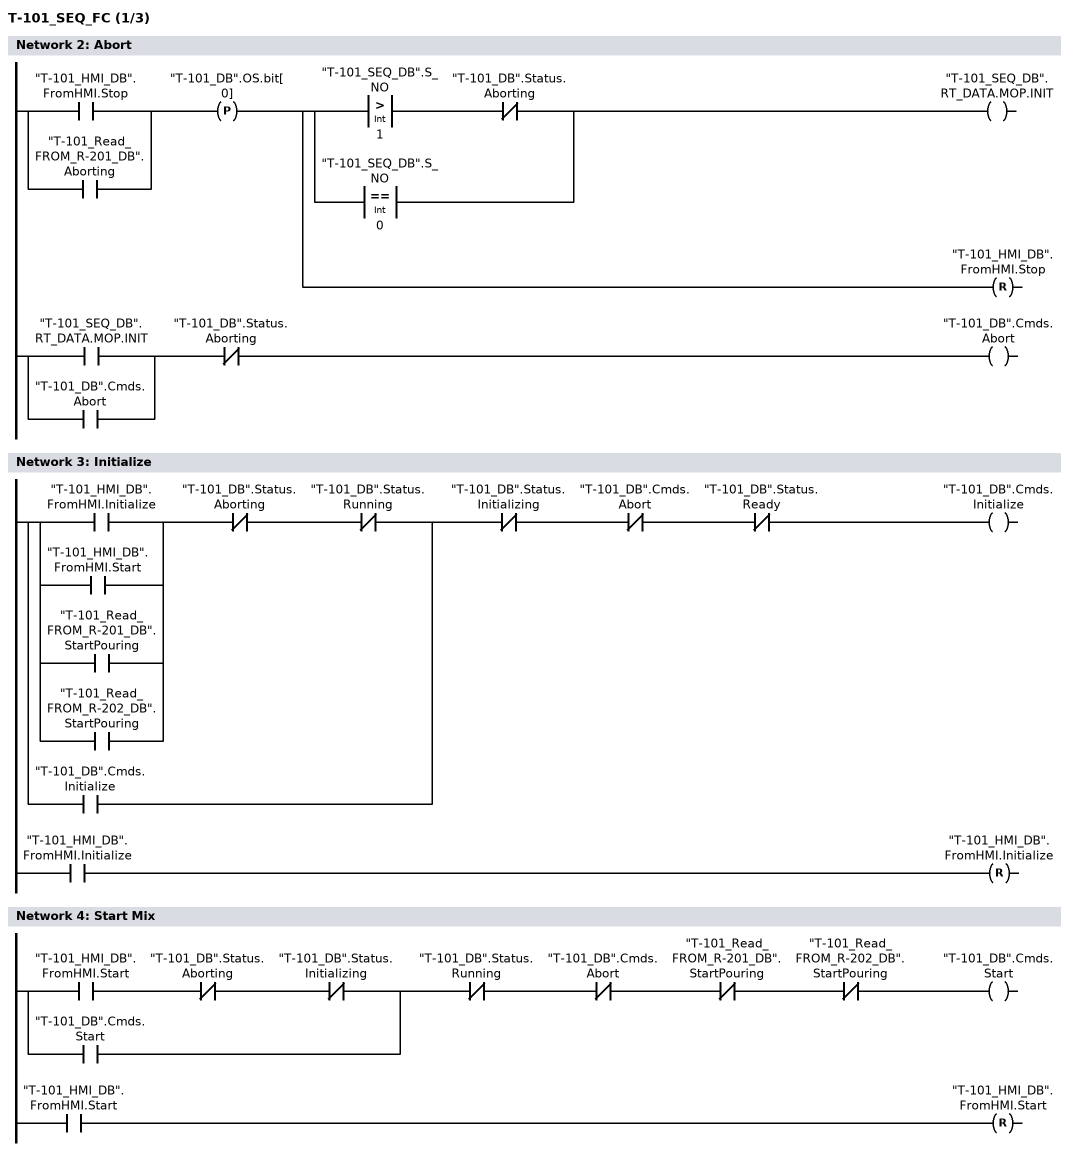
   RUNG wire#powerrail
      Contact( "T-101_HMI_DB".FromHMI.Stop )
      wire#w1
      P_Trig( "T-101_DB".OS.bit[0] )
      wire#w2
      { S7_Templates := "SrcType := Int" } GT_Contact(in1 := "T-101_SEQ_DB".S_NO, in2 := 1)
      I_Contact( "T-101_DB".Status.Aborting )
      wire#w3
      Coil( "T-101_SEQ_DB".RT_DATA.MOP.INIT )
   END_RUNG
   RUNG wire#powerrail
      Contact( "T-101_Read_FROM_R-201_DB".Aborting )
   END_RUNG wire#w1
   RUNG wire#w2
      { S7_Templates := "SrcType := Int" } EQ_Contact(in1 := "T-101_SEQ_DB".S_NO, in2 := 0)
   END_RUNG wire#w3
   RUNG wire#w2
      R_Coil( "T-101_HMI_DB".FromHMI.Stop )
   END_RUNG
   RUNG wire#powerrail
      Contact( "T-101_SEQ_DB".RT_DATA.MOP.INIT )
      wire#w4
      I_Contact( "T-101_DB".Status.Aborting )
      Coil( "T-101_DB".Cmds.Abort )
   END_RUNG
   RUNG wire#powerrail
      Contact( "T-101_DB".Cmds.Abort )
   END_RUNG wire#w4
   // the same network as SCL:
   #_w1 := "T-101_HMI_DB".FromHMI.Stop OR "T-101_Read_FROM_R-201_DB".Aborting;
   #_w2 := #_w1 AND NOT "T-101_DB".OS.bit[0];   // rising edge
   "T-101_DB".OS.bit[0] := #_w1;
   "T-101_SEQ_DB".RT_DATA.MOP.INIT := #_w2 AND ((("T-101_SEQ_DB".S_NO > 1) AND NOT "T-101_DB".Status.Aborting) OR ("T-101_SEQ_DB".S_NO = 0));
   IF #_w2 THEN "T-101_HMI_DB".FromHMI.Stop := FALSE; END_IF;
   "T-101_DB".Cmds.Abort := ("T-101_SEQ_DB".RT_DATA.MOP.INIT OR "T-101_DB".Cmds.Abort) AND NOT "T-101_DB".Status.Aborting;
END_REGION

REGION Network 3: Initialize
   RUNG wire#powerrail
      Contact( "T-101_HMI_DB".FromHMI.Initialize )
      wire#w1
      I_Contact( "T-101_DB".Status.Aborting )
      I_Contact( "T-101_DB".Status.Running )
      wire#w2
      I_Contact( "T-101_DB".Status.Initializing )
      I_Contact( "T-101_DB".Cmds.Abort )
      I_Contact( "T-101_DB".Status.Ready )
      Coil( "T-101_DB".Cmds.Initialize )
   END_RUNG
   RUNG wire#powerrail
      Contact( "T-101_HMI_DB".FromHMI.Start )
   END_RUNG wire#w1
   RUNG wire#powerrail
      Contact( "T-101_Read_FROM_R-201_DB".StartPouring )
   END_RUNG wire#w1
   RUNG wire#powerrail
      Contact( "T-101_Read_FROM_R-202_DB".StartPouring )
   END_RUNG wire#w1
   RUNG wire#powerrail
      Contact( "T-101_DB".Cmds.Initialize )
   END_RUNG wire#w2
   RUNG wire#powerrail
      Contact( "T-101_HMI_DB".FromHMI.Initialize )
      R_Coil( "T-101_HMI_DB".FromHMI.Initialize )
   END_RUNG
   // the same network as SCL:
   "T-101_DB".Cmds.Initialize := ((("T-101_HMI_DB".FromHMI.Initialize OR "T-101_HMI_DB".FromHMI.Start OR "T-101_Read_FROM_R-201_DB".StartPouring OR "T-101_Read_FROM_R-202_DB".StartPouring) AND NOT "T-101_DB".Status.Aborting AND NOT "T-101_DB".Status.Running) OR "T-101_DB".Cmds.Initialize) AND NOT "T-101_DB".Status.Initializing AND NOT "T-101_DB".Cmds.Abort AND NOT "T-101_DB".Status.Ready;
   IF "T-101_HMI_DB".FromHMI.Initialize THEN "T-101_HMI_DB".FromHMI.Initialize := FALSE; END_IF;
END_REGION

REGION Network 4: Start Mix
   RUNG wire#powerrail
      Contact( "T-101_HMI_DB".FromHMI.Start )
      I_Contact( "T-101_DB".Status.Aborting )
      I_Contact( "T-101_DB".Status.Initializing )
      wire#w1
      I_Contact( "T-101_DB".Status.Running )
      I_Contact( "T-101_DB".Cmds.Abort )
      I_Contact( "T-101_Read_FROM_R-201_DB".StartPouring )
      I_Contact( "T-101_Read_FROM_R-202_DB".StartPouring )
      Coil( "T-101_DB".Cmds.Start )
   END_RUNG
   RUNG wire#powerrail
      Contact( "T-101_DB".Cmds.Start )
   END_RUNG wire#w1
   RUNG wire#powerrail
      Contact( "T-101_HMI_DB".FromHMI.Start )
      R_Coil( "T-101_HMI_DB".FromHMI.Start )
   END_RUNG
   // the same network as SCL:
   "T-101_DB".Cmds.Start := (("T-101_HMI_DB".FromHMI.Start AND NOT "T-101_DB".Status.Aborting AND NOT "T-101_DB".Status.Initializing) OR "T-101_DB".Cmds.Start) AND NOT "T-101_DB".Status.Running AND NOT "T-101_DB".Cmds.Abort AND NOT "T-101_Read_FROM_R-201_DB".StartPouring AND NOT "T-101_Read_FROM_R-202_DB".StartPouring;
   IF "T-101_HMI_DB".FromHMI.Start THEN "T-101_HMI_DB".FromHMI.Start := FALSE; END_IF;
END_REGION

REGION Network 5: Procedure Selected
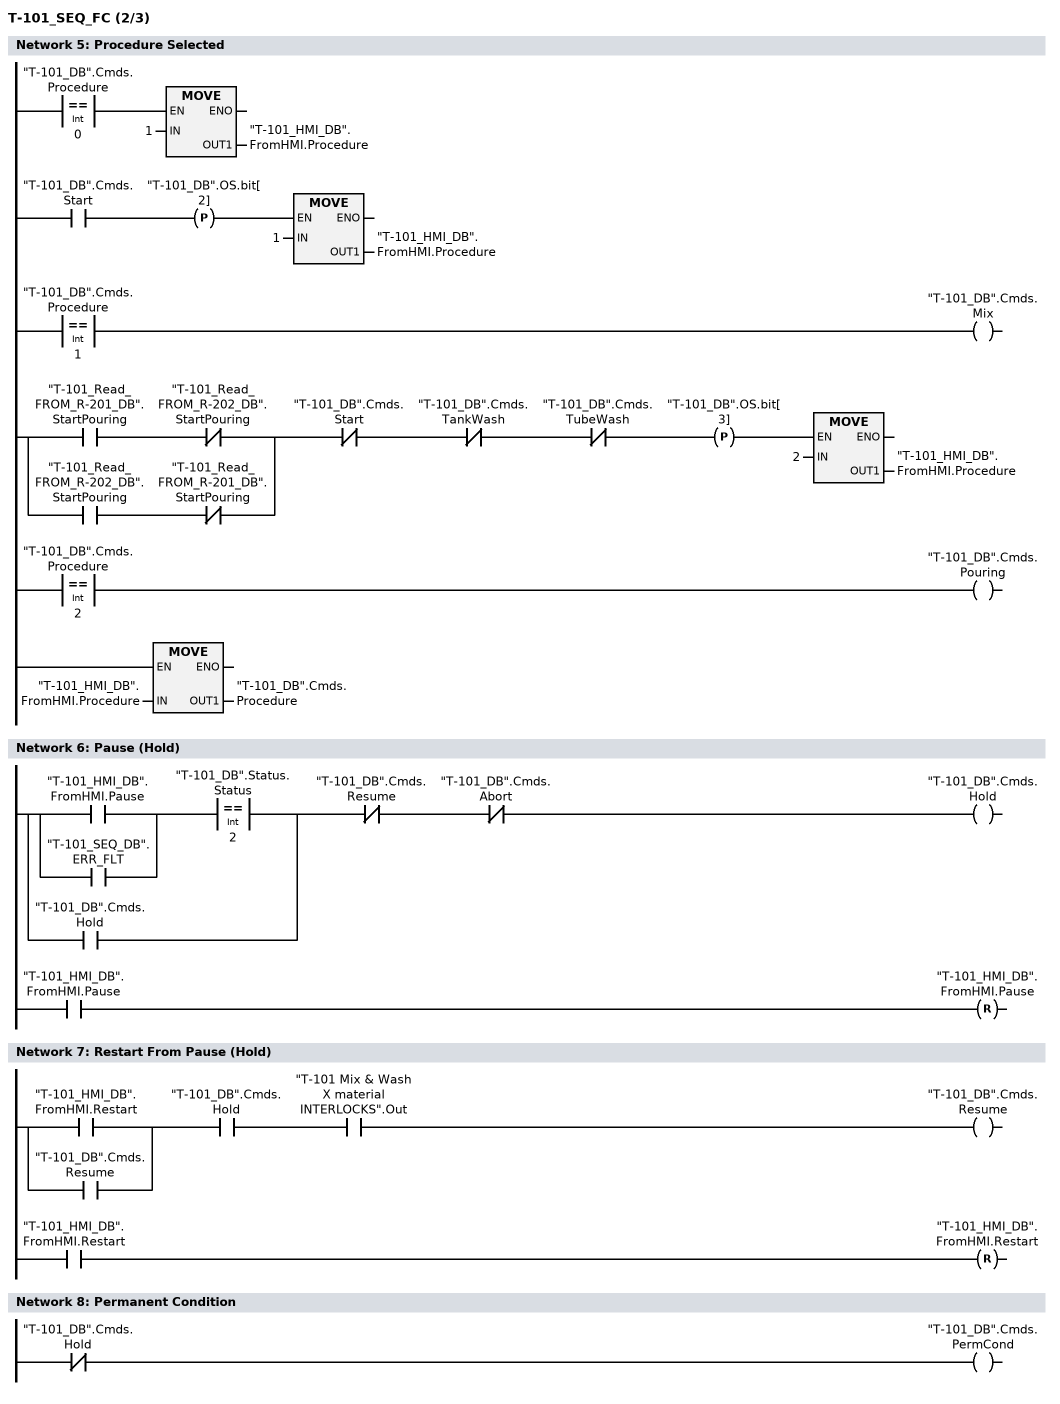
   RUNG wire#powerrail
      { S7_Templates := "SrcType := Int" } EQ_Contact(in1 := "T-101_DB".Cmds.Procedure, in2 := 0)
      Move(in := 1, out1 => "T-101_HMI_DB".FromHMI.Procedure)
   END_RUNG
   RUNG wire#powerrail
      Contact( "T-101_DB".Cmds.Start )
      P_Trig( "T-101_DB".OS.bit[2] )
      Move(in := 1, out1 => "T-101_HMI_DB".FromHMI.Procedure)
   END_RUNG
   RUNG wire#powerrail
      { S7_Templates := "SrcType := Int" } EQ_Contact(in1 := "T-101_DB".Cmds.Procedure, in2 := 1)
      Coil( "T-101_DB".Cmds.Mix )
   END_RUNG
   RUNG wire#powerrail
      Contact( "T-101_Read_FROM_R-201_DB".StartPouring )
      I_Contact( "T-101_Read_FROM_R-202_DB".StartPouring )
      wire#w1
      I_Contact( "T-101_DB".Cmds.Start )
      I_Contact( "T-101_DB".Cmds.TankWash )
      I_Contact( "T-101_DB".Cmds.TubeWash )
      P_Trig( "T-101_DB".OS.bit[3] )
      Move(in := 2, out1 => "T-101_HMI_DB".FromHMI.Procedure)
   END_RUNG
   RUNG wire#powerrail
      Contact( "T-101_Read_FROM_R-202_DB".StartPouring )
      I_Contact( "T-101_Read_FROM_R-201_DB".StartPouring )
   END_RUNG wire#w1
   RUNG wire#powerrail
      { S7_Templates := "SrcType := Int" } EQ_Contact(in1 := "T-101_DB".Cmds.Procedure, in2 := 2)
      Coil( "T-101_DB".Cmds.Pouring )
   END_RUNG
   RUNG wire#powerrail
      Move(in := "T-101_HMI_DB".FromHMI.Procedure, out1 => "T-101_DB".Cmds.Procedure)
   END_RUNG
   // the same network as SCL:
   IF "T-101_DB".Cmds.Procedure = 0 THEN "T-101_HMI_DB".FromHMI.Procedure := 1; END_IF;
   #_w1 := "T-101_DB".Cmds.Start AND NOT "T-101_DB".OS.bit[2];   // rising edge
   "T-101_DB".OS.bit[2] := "T-101_DB".Cmds.Start;
   IF #_w1 THEN "T-101_HMI_DB".FromHMI.Procedure := 1; END_IF;
   "T-101_DB".Cmds.Mix := "T-101_DB".Cmds.Procedure = 1;
   #_w2 := (("T-101_Read_FROM_R-201_DB".StartPouring AND NOT "T-101_Read_FROM_R-202_DB".StartPouring) OR ("T-101_Read_FROM_R-202_DB".StartPouring AND NOT "T-101_Read_FROM_R-201_DB".StartPouring)) AND NOT "T-101_DB".Cmds.Start AND NOT "T-101_DB".Cmds.TankWash AND NOT "T-101_DB".Cmds.TubeWash;
   #_w3 := #_w2 AND NOT "T-101_DB".OS.bit[3];   // rising edge
   "T-101_DB".OS.bit[3] := #_w2;
   IF #_w3 THEN "T-101_HMI_DB".FromHMI.Procedure := 2; END_IF;
   "T-101_DB".Cmds.Pouring := "T-101_DB".Cmds.Procedure = 2;
   "T-101_DB".Cmds.Procedure := "T-101_HMI_DB".FromHMI.Procedure;
END_REGION

REGION Network 6: Pause (Hold)
   RUNG wire#powerrail
      Contact( "T-101_HMI_DB".FromHMI.Pause )
      wire#w1
      { S7_Templates := "SrcType := Int" } EQ_Contact(in1 := "T-101_DB".Status.Status, in2 := 2)
      wire#w2
      I_Contact( "T-101_DB".Cmds.Resume )
      I_Contact( "T-101_DB".Cmds.Abort )
      Coil( "T-101_DB".Cmds.Hold )
   END_RUNG
   RUNG wire#powerrail
      Contact( "T-101_SEQ_DB".ERR_FLT )
   END_RUNG wire#w1
   RUNG wire#powerrail
      Contact( "T-101_DB".Cmds.Hold )
   END_RUNG wire#w2
   RUNG wire#powerrail
      Contact( "T-101_HMI_DB".FromHMI.Pause )
      R_Coil( "T-101_HMI_DB".FromHMI.Pause )
   END_RUNG
   // the same network as SCL:
   "T-101_DB".Cmds.Hold := ((("T-101_HMI_DB".FromHMI.Pause OR "T-101_SEQ_DB".ERR_FLT) AND ("T-101_DB".Status.Status = 2)) OR "T-101_DB".Cmds.Hold) AND NOT "T-101_DB".Cmds.Resume AND NOT "T-101_DB".Cmds.Abort;
   IF "T-101_HMI_DB".FromHMI.Pause THEN "T-101_HMI_DB".FromHMI.Pause := FALSE; END_IF;
END_REGION

REGION Network 7: Restart From Pause (Hold)
   RUNG wire#powerrail
      Contact( "T-101_HMI_DB".FromHMI.Restart )
      wire#w1
      Contact( "T-101_DB".Cmds.Hold )
      Contact( "T-101 Mix & Wash X material INTERLOCKS".Out )
      Coil( "T-101_DB".Cmds.Resume )
   END_RUNG
   RUNG wire#powerrail
      Contact( "T-101_DB".Cmds.Resume )
   END_RUNG wire#w1
   RUNG wire#powerrail
      Contact( "T-101_HMI_DB".FromHMI.Restart )
      R_Coil( "T-101_HMI_DB".FromHMI.Restart )
   END_RUNG
   // the same network as SCL:
   "T-101_DB".Cmds.Resume := ("T-101_HMI_DB".FromHMI.Restart OR "T-101_DB".Cmds.Resume) AND "T-101_DB".Cmds.Hold AND "T-101 Mix & Wash X material INTERLOCKS".Out;
   IF "T-101_HMI_DB".FromHMI.Restart THEN "T-101_HMI_DB".FromHMI.Restart := FALSE; END_IF;
END_REGION

REGION Network 8: Permanent Condition
   RUNG wire#powerrail
      I_Contact( "T-101_DB".Cmds.Hold )
      Coil( "T-101_DB".Cmds.PermCond )
   END_RUNG
   // the same network as SCL:
   "T-101_DB".Cmds.PermCond := NOT "T-101_DB".Cmds.Hold;
END_REGION

REGION Network 9: Tank Wash
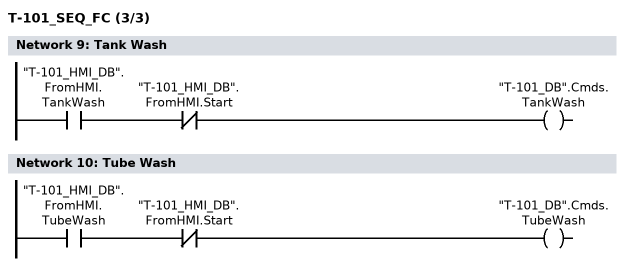
   RUNG wire#powerrail
      Contact( "T-101_HMI_DB".FromHMI.TankWash )
      I_Contact( "T-101_HMI_DB".FromHMI.Start )
      Coil( "T-101_DB".Cmds.TankWash )
   END_RUNG
   // the same network as SCL:
   "T-101_DB".Cmds.TankWash := "T-101_HMI_DB".FromHMI.TankWash AND NOT "T-101_HMI_DB".FromHMI.Start;
END_REGION

REGION Network 10: Tube Wash
   RUNG wire#powerrail
      Contact( "T-101_HMI_DB".FromHMI.TubeWash )
      I_Contact( "T-101_HMI_DB".FromHMI.Start )
      Coil( "T-101_DB".Cmds.TubeWash )
   END_RUNG
   // the same network as SCL:
   "T-101_DB".Cmds.TubeWash := "T-101_HMI_DB".FromHMI.TubeWash AND NOT "T-101_HMI_DB".FromHMI.Start;
END_REGION

REGION Network 11 (SCL): Sequence Status
   IF "T-101_SEQ_DB".S_NO = 1 THEN
       "T-101_DB".Status.Status := 1; //Idle
   ELSIF ("T-101_SEQ_DB".S_NO > 1 AND "T-101_SEQ_DB".S_NO < 150) AND NOT "T-101_SEQ_DB".ERR_FLT AND NOT "T-101_DB".Cmds.Hold THEN
       "T-101_DB".Status.Status := 2; //Running
   ELSIF "T-101_SEQ_DB".S_NO >= 151 AND "T-101_SEQ_DB".S_NO <= 160 AND NOT "T-101_SEQ_DB".ERR_FLT THEN
       "T-101_DB".Status.Status := 3; // Stopping
   ELSIF "T-101_SEQ_DB".ERR_FLT AND ("T-101_SEQ_DB".S_NO > 1 AND "T-101_SEQ_DB".S_NO < 150) THEN
       "T-101_DB".Status.Status := 4; // Held
   ELSIF "T-101_SEQ_DB".ERR_FLT AND ("T-101_SEQ_DB".S_NO > 1 AND "T-101_SEQ_DB".S_NO < 150) AND "T-101_Aux_DB"."Bool".TOff THEN
       "T-101_DB".Status.Status := 5; // Holding
   ELSE
       "T-101_DB".Status.Status := 6; // Unknown
   END_IF;

   "T-101_DB".Status.Running := ("T-101_SEQ_DB".S_NO > 3 AND "T-101_SEQ_DB".S_NO <= 150);
   "T-101_DB".Status.Initializing := ("T-101_SEQ_DB".S_NO >= 141 AND "T-101_SEQ_DB".S_NO <= 150);
   //"T-101_DB".Status.Aborting := ("T-101_SEQ_DB".S_NO >= 151 AND "T-101_SEQ_DB".S_NO <= 160);

   //Enable/Disable HMI Start/Stop Button
   "T-101_HMI_DB".ToHMI.EnStopButton := ("T-101_DB".Status.Status > 1) OR "T-101_DB".Status.Step = 0; //Enable HMI Stop Button
   "T-101_HMI_DB".ToHMI.EnStartButton := "T-101_DB".Status.Status = 1; //Idle
   "T-101_HMI_DB".ToHMI.EnPauseButton := "T-101_DB".Status.Status = 2; //Enable Pause Button
   "T-101_HMI_DB".ToHMI.EnRestartButton :=  "T-101_DB".Status.Status = 4 ; //Enable Restart Button

   //****Interlock Activated
   "T-101_HMI_DB".ToHMI.InterlockActivated := "T-101 Mix & Wash X material INTERLOCKS".Out;
END_REGION

REGION Network 12 (SCL): Sequence Step
   "T-101_DB".Status.Step := "T-101_SEQ_DB".S_NO;
END_REGION

REGION Network 13 (SCL): Sequence state (Procedure running)
   IF "T-101_SEQ_DB".S_NO = 3 OR "T-101_SEQ_DB".S_NO = 4 THEN
       "T-101_DB".Status.State := 1; //Ready
   ELSIF "T-101_SEQ_DB".S_NO >= 21 AND "T-101_SEQ_DB".S_NO <= 60 THEN
       "T-101_DB".Status.State := 2; //Mixing 
   ELSIF "T-101_SEQ_DB".S_NO >= 61 AND "T-101_SEQ_DB".S_NO <= 80 THEN
       "T-101_DB".Status.State := 3; //Pouring
   ELSIF "T-101_SEQ_DB".S_NO >= 141 AND "T-101_SEQ_DB".S_NO <= 150 THEN
       "T-101_DB".Status.State := 4; //Initializing
   ELSIF "T-101_SEQ_DB".S_NO >= 151 AND "T-101_SEQ_DB".S_NO <= 160 THEN
       "T-101_DB".Status.State := 5; //Aborting
   ELSE
       "T-101_DB".Status.State := 0;
   END_IF;
END_REGION

REGION Network 14: Sequence State
END_REGION
END_FUNCTION

FUNCTION "T-101_FC_Outputs" : Void   // FC81, SCL
{ S7_Optimized_Access := 'TRUE' }
VERSION : 0.1
   VAR_TEMP
      Pump_A : Struct
         Cond_01 : Bool;   // Condition 01
         Cond_02 : Bool;
         Cond_03 : Bool;   // Condition 03
      END_STRUCT;
      Pump_B : Struct
         Cond_01 : Bool;   // Condition 01
         Cond_02 : Bool;   // Condition 02
         Cond_03 : Bool;   // Condition 03
      END_STRUCT;
      XV : Struct
         "1011" : Bool;
         "1041" : Bool;
         "1013" : Bool;
      END_STRUCT;
      RouteOpened : Bool;
      PumpsOff : Bool;
      Recirculating : Bool;
   END_VAR
BEGIN
   //****** Equipmens Activation*******
   //
   //**************************************************************
   //

   //
   //IF "AlwaysFALSE" THEN
       //***********************************************Tank Outlet Valve**********************************************************************
       IF  "XV-1011_DB".Mode=0 THEN
           "T-101_DB".Equipments.Valves."XV-1011".CmdOn := "T-101_DB".Equipments.Valves."XV-1011".Enable AND NOT "T-101_DB".Cmds.Hold;
           //Delay Off To avoid Overpressure the Lines
           #XV."1011" := "T-101_DB".Equipments.Valves."XV-1011".CmdOn;
           "T-101_Aux_DB".Timer."XV-1011".TOF(IN := #XV."1011",
                                              PT := "T-101_Aux_DB".Constants.CmdDelay);
           //Command to the Valve
           IF "T-101_Aux_DB".Timer."XV-1011".Q THEN
               "XV-1011_DB".CMD := 2;
           ELSE
               "XV-1011_DB".CMD := 1;
           END_IF;
           "T-101_DB".Equipments.Valves."XV-1011".TurningOff := NOT "T-101_DB".Equipments.Valves."XV-1011".CmdOn AND "T-101_Aux_DB".Timer."XV-1011".Q;
       END_IF;
       //***********************************************Tank Inlet Valve**********************************************************************
       IF  "XV-1041_DB".Mode = 0 THEN
           "T-101_DB".Equipments.Valves."XV-1041".CmdOn := "T-101_DB".Equipments.Valves."XV-1041".Enable AND NOT "T-101_DB".Cmds.Hold;
           //Delay Off To avoid Overpressure the Lines
           #XV."1041" := "T-101_DB".Equipments.Valves."XV-1041".CmdOn;
           "T-101_Aux_DB".Timer."XV-1041".TOF(IN := #XV."1041",
                                              PT := "T-101_Aux_DB".Constants.CmdDelay);
           //Command to the Valve
           IF "T-101_Aux_DB".Timer."XV-1041".Q THEN
               "XV-1041_DB".CMD := 2;
           ELSE
               "XV-1041_DB".CMD := 1;
           END_IF;
           "T-101_DB".Equipments.Valves."XV-1041".TurningOff := NOT "T-101_DB".Equipments.Valves."XV-1041".CmdOn AND "T-101_Aux_DB".Timer."XV-1041".Q;
       END_IF;
       //***********************************************Tank Transfer Valve**********************************************************************
       IF  "XV-1013_DB".Mode = 0 THEN
           "T-101_DB".Equipments.Valves."XV-1013".CmdOn := "T-101_DB".Equipments.Valves."XV-1013".Enable AND NOT "T-101_DB".Cmds.Hold;
           //Delay Off To avoid Overpressure the Lines
           #XV."1013" := "T-101_DB".Equipments.Valves."XV-1013".CmdOn;
           "T-101_Aux_DB".Timer."XV-1013".TOF(IN := #XV."1013",
                                              PT := "T-101_Aux_DB".Constants.CmdDelay);
           //Command to the Valve
           IF "T-101_Aux_DB".Timer."XV-1013".Q THEN
               "XV-1013_DB".CMD := 2;
           ELSE
               "XV-1013_DB".CMD := 1;
           END_IF;
           "T-101_DB".Equipments.Valves."XV-1013".TurningOff := NOT "T-101_DB".Equipments.Valves."XV-1013".CmdOn AND "T-101_Aux_DB".Timer."XV-1013".Q;
       END_IF;
      // IF NOT "TestDB".DesablePmps_T101 THEN
           //***********************************************Feed Water Pump A**********************************************************************
           // Condition to CmdOn "On Command" 
           IF  "P-101A_DB".Config.HMI.Enable_HMI_Controls=1 THEN
               #Pump_A.Cond_01 := "T-101_DB".Equipments.Pumps."P-101A".Enable AND ("T-101_DB".PmpSel."P-101AB" = 1 OR "T-101_DB".PmpSel."P-101AB" = 3);
               #Pump_A.Cond_02 := "T-101_Write_TO_R-201_DB".RouteOpened AND "T-101_Read_FROM_R-201_DB".RouteOpened OR ("T-101_Write_TO_R-202_DB".RouteOpened AND "T-101_Read_FROM_R-202_DB".RouteOpened); //Route Open to sent to the Reactor
               #Pump_A.Cond_03 := "XV-1011_DB".OS AND "XV-1013_DB".CS; //Route open to Recirculate
               "T-101_DB".Equipments.Pumps."P-101A".CmdOn := #Pump_A.Cond_01 AND (#Pump_A.Cond_02 OR #Pump_A.Cond_03) AND NOT "T-101_DB".Cmds.Hold;
               IF "T-101_DB".Equipments.Pumps."P-101A".CmdOn THEN
                   "P-101A_DB".Stop_CMD := False;
                   "P-101A_DB".Start_CMD := true;
                   "P-101A_DB".ON := TRUE;
                   "P-101A_DB".OFF := FALSE;
               ELSE
                   "P-101A_DB".Stop_CMD := true;
                   "P-101A_DB".Start_CMD :=false;
                   "P-101A_DB".ON := FALSE;
                   "P-101A_DB".OFF := TRUE;
               END_IF;
           END_IF;
           //***********************************************Feed Water Pump B**********************************************************************
           // Condition to CmdOn "On Command" 
           IF  "P-101B_DB".Config.HMI.Enable_HMI_Controls = 1 THEN
               #Pump_B.Cond_01 := "T-101_DB".Equipments.Pumps."P-101B".Enable AND ("T-101_DB".PmpSel."P-101AB" = 2 OR "T-101_DB".PmpSel."P-101AB" = 3);
               #Pump_B.Cond_02 := "T-101_Write_TO_R-201_DB".RouteOpened AND "T-101_Read_FROM_R-201_DB".RouteOpened  OR ("T-101_Write_TO_R-202_DB".RouteOpened AND "T-101_Read_FROM_R-202_DB".RouteOpened); //Route Open to sent to the Reactor
               #Pump_B.Cond_03 := "XV-1011_DB".OS AND "XV-1013_DB".CS; //Route open to Recirculate
               "T-101_DB".Equipments.Pumps."P-101B".CmdOn := #Pump_B.Cond_01 AND (#Pump_B.Cond_02 OR #Pump_B.Cond_03) AND NOT "T-101_DB".Cmds.Hold;
               IF "T-101_DB".Equipments.Pumps."P-101B".CmdOn THEN
                   "P-101B_DB".Stop_CMD := False;
                   "P-101B_DB".Start_CMD := true;
                   "P-101B_DB".ON := TRUE;
                   "P-101B_DB".OFF := FALSE;
               ELSE
                   "P-101B_DB".Stop_CMD := True;
                   "P-101B_DB".Start_CMD := False;
                   "P-101B_DB".ON := FALSE;
                   "P-101B_DB".OFF := TRUE;
               END_IF;
           END_IF;
       //END_IF;
           //***********************************************Mixer***********************************************************************
           IF "VFD-T101A_DB".HMI.Controls.Mode = 2 THEN
               "T-101_DB".Equipments.VFD."VFD-1011".CmdOn := "T-101_DB".Equipments.VFD."VFD-1011".Enable AND NOT "T-101_DB".Cmds.Hold;
               IF "T-101_DB".Equipments.VFD."VFD-1011".CmdOn THEN
                   "VFD-T101A_DB".PLCCommand := TRUE;
               ELSE
                   "VFD-T101A_DB".PLCCommand := FALSE;
               END_IF;
           END_IF;
       //END_IF;


   //END_IF;

   //***************Interlocks to R-201***************//
   //*****Recirculating*****//
   #Recirculating := ("P-101A_DB".CF OR "P-101B_DB".CF) AND ("XV-1011_DB".OS AND "XV-1013_DB".CS) AND ("FT-1011_DB".SAI > 0.2);

   "T-101_Write_TO_R-201_DB".Recirculating :=    #Recirculating;
   "T-101_Write_TO_R-202_DB".Recirculating :=    #Recirculating;
   //****Route open to R-201*****//
           #RouteOpened := "XV-1011_DB".OS AND "XV-1013_DB".OS;

   "T-101_Write_TO_R-201_DB".RouteOpened :=   #RouteOpened ;
   "T-101_Write_TO_R-202_DB".RouteOpened := #RouteOpened;
   //*****Pumps OFF*****//
   #PumpsOff := NOT "P-101A_DB".CF AND NOT "P-101B_DB".CF AND ("PT-101A_DB".SAI < 0.8 AND "PT-101B_DB".SAI < 0.8);

   "T-101_Write_TO_R-201_DB".PupmsOFF :=  #PumpsOff ;
   "T-101_Write_TO_R-202_DB".PupmsOFF :=  #PumpsOff ;

           //********************Tank Internal Status*********************************
   "T-101_DB".Status.PouringRunning := ("T-101_DB".Status.Step = 61 OR "T-101_DB".Status.Step = 62 OR "T-101_DB".Status.Step = 63) AND (#RouteOpened AND NOT #PumpsOff);

   //***************Interlocks to T-104***************//
   "T-101_Write_TO_T-104_DB".ReqWaterToMix := "XV-1041_DB".OS AND "T-101_DB".ExchangeCmds.Send.ReqWater;
   "T-101_Write_TO_T-104_DB".StopReqWaterToMix := "T-101_DB".ExchangeCmds.Send.StopReqWater;

   //***************Valves Status***************//
   "T-101_Aux_DB"."Bool".TOff := "T-101_DB".Equipments.Valves."XV-1011".TurningOff OR "T-101_DB".Equipments.Valves."XV-1041".TurningOff OR "T-101_DB".Equipments.Valves."XV-1013".TurningOff;
   //***************Timer***************//
   "T-101_Aux_DB"."Bool".MinMixT_Enab := "T-101_DB".Status.Step = 27 AND "VFD-T101A_DB".RUN_FEEDBACK AND "VFD-T101A_DB".SPEED_FEEDBACK > 500;
   "T-101_Aux_DB"."Bool".MinMixT_Reset := "T-101_DB".Cmds.Abort OR "T-101_DB".Status.Step = 1;
END_FUNCTION

// folder: State MACHINE/1)Tanks/Tank T-101 (X)/T-101 <---> R-201

FUNCTION "T-101_Signals_FROM_R-201" : Void   // FC66, LAD
{ S7_Optimized_Access := 'TRUE' }
VERSION : 0.1
BEGIN

REGION Network 1: Start Pouring Sequence
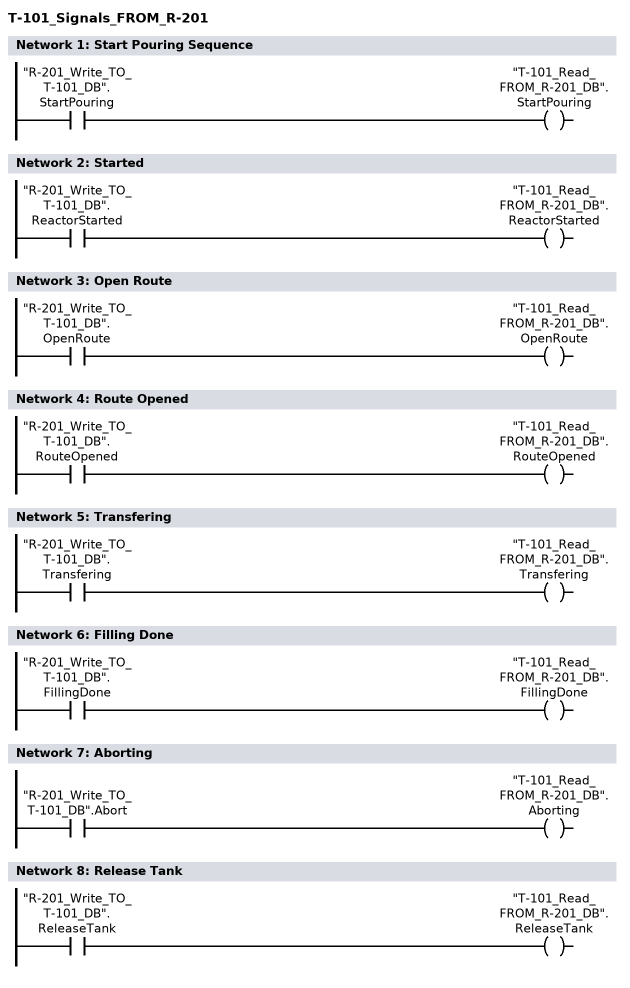
   RUNG wire#powerrail
      Contact( "R-201_Write_TO_T-101_DB".StartPouring )
      Coil( "T-101_Read_FROM_R-201_DB".StartPouring )
   END_RUNG
   // the same network as SCL:
   "T-101_Read_FROM_R-201_DB".StartPouring := "R-201_Write_TO_T-101_DB".StartPouring;
END_REGION

REGION Network 2: Started
   RUNG wire#powerrail
      Contact( "R-201_Write_TO_T-101_DB".ReactorStarted )
      Coil( "T-101_Read_FROM_R-201_DB".ReactorStarted )
   END_RUNG
   // the same network as SCL:
   "T-101_Read_FROM_R-201_DB".ReactorStarted := "R-201_Write_TO_T-101_DB".ReactorStarted;
END_REGION

REGION Network 3: Open Route
   RUNG wire#powerrail
      Contact( "R-201_Write_TO_T-101_DB".OpenRoute )
      Coil( "T-101_Read_FROM_R-201_DB".OpenRoute )
   END_RUNG
   // the same network as SCL:
   "T-101_Read_FROM_R-201_DB".OpenRoute := "R-201_Write_TO_T-101_DB".OpenRoute;
END_REGION

REGION Network 4: Route Opened
   RUNG wire#powerrail
      Contact( "R-201_Write_TO_T-101_DB".RouteOpened )
      Coil( "T-101_Read_FROM_R-201_DB".RouteOpened )
   END_RUNG
   // the same network as SCL:
   "T-101_Read_FROM_R-201_DB".RouteOpened := "R-201_Write_TO_T-101_DB".RouteOpened;
END_REGION

REGION Network 5: Transfering
   RUNG wire#powerrail
      Contact( "R-201_Write_TO_T-101_DB".Transfering )
      Coil( "T-101_Read_FROM_R-201_DB".Transfering )
   END_RUNG
   // the same network as SCL:
   "T-101_Read_FROM_R-201_DB".Transfering := "R-201_Write_TO_T-101_DB".Transfering;
END_REGION

REGION Network 6: Filling Done
   RUNG wire#powerrail
      Contact( "R-201_Write_TO_T-101_DB".FillingDone )
      Coil( "T-101_Read_FROM_R-201_DB".FillingDone )
   END_RUNG
   // the same network as SCL:
   "T-101_Read_FROM_R-201_DB".FillingDone := "R-201_Write_TO_T-101_DB".FillingDone;
END_REGION

REGION Network 7: Aborting
   RUNG wire#powerrail
      Contact( "R-201_Write_TO_T-101_DB".Abort )
      Coil( "T-101_Read_FROM_R-201_DB".Aborting )
   END_RUNG
   // the same network as SCL:
   "T-101_Read_FROM_R-201_DB".Aborting := "R-201_Write_TO_T-101_DB".Abort;
END_REGION

REGION Network 8: Release Tank
   RUNG wire#powerrail
      Contact( "R-201_Write_TO_T-101_DB".ReleaseTank )
      Coil( "T-101_Read_FROM_R-201_DB".ReleaseTank )
   END_RUNG
   // the same network as SCL:
   "T-101_Read_FROM_R-201_DB".ReleaseTank := "R-201_Write_TO_T-101_DB".ReleaseTank;
END_REGION
END_FUNCTION

// folder: State MACHINE/1)Tanks/Tank T-101 (X)/T-101 <---> R-202

FUNCTION "T-101_Signals_FROM_R-202" : Void   // FC65, LAD
{ S7_Optimized_Access := 'TRUE' }
VERSION : 0.1
BEGIN

REGION Network 1: Start Pouring Sequence
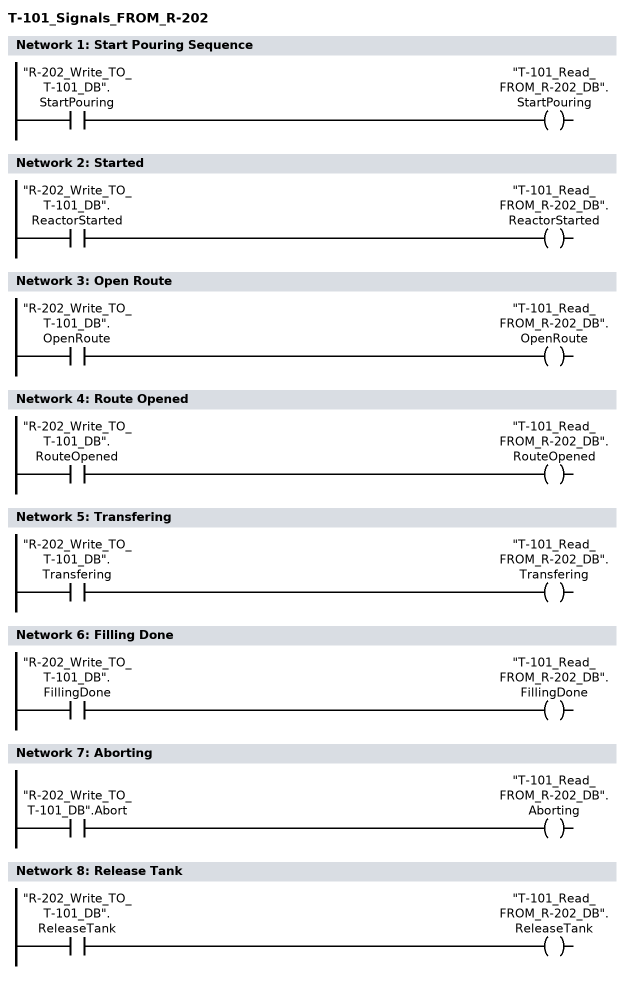
   RUNG wire#powerrail
      Contact( "R-202_Write_TO_T-101_DB".StartPouring )
      Coil( "T-101_Read_FROM_R-202_DB".StartPouring )
   END_RUNG
   // the same network as SCL:
   "T-101_Read_FROM_R-202_DB".StartPouring := "R-202_Write_TO_T-101_DB".StartPouring;
END_REGION

REGION Network 2: Started
   RUNG wire#powerrail
      Contact( "R-202_Write_TO_T-101_DB".ReactorStarted )
      Coil( "T-101_Read_FROM_R-202_DB".ReactorStarted )
   END_RUNG
   // the same network as SCL:
   "T-101_Read_FROM_R-202_DB".ReactorStarted := "R-202_Write_TO_T-101_DB".ReactorStarted;
END_REGION

REGION Network 3: Open Route
   RUNG wire#powerrail
      Contact( "R-202_Write_TO_T-101_DB".OpenRoute )
      Coil( "T-101_Read_FROM_R-202_DB".OpenRoute )
   END_RUNG
   // the same network as SCL:
   "T-101_Read_FROM_R-202_DB".OpenRoute := "R-202_Write_TO_T-101_DB".OpenRoute;
END_REGION

REGION Network 4: Route Opened
   RUNG wire#powerrail
      Contact( "R-202_Write_TO_T-101_DB".RouteOpened )
      Coil( "T-101_Read_FROM_R-202_DB".RouteOpened )
   END_RUNG
   // the same network as SCL:
   "T-101_Read_FROM_R-202_DB".RouteOpened := "R-202_Write_TO_T-101_DB".RouteOpened;
END_REGION

REGION Network 5: Transfering
   RUNG wire#powerrail
      Contact( "R-202_Write_TO_T-101_DB".Transfering )
      Coil( "T-101_Read_FROM_R-202_DB".Transfering )
   END_RUNG
   // the same network as SCL:
   "T-101_Read_FROM_R-202_DB".Transfering := "R-202_Write_TO_T-101_DB".Transfering;
END_REGION

REGION Network 6: Filling Done
   RUNG wire#powerrail
      Contact( "R-202_Write_TO_T-101_DB".FillingDone )
      Coil( "T-101_Read_FROM_R-202_DB".FillingDone )
   END_RUNG
   // the same network as SCL:
   "T-101_Read_FROM_R-202_DB".FillingDone := "R-202_Write_TO_T-101_DB".FillingDone;
END_REGION

REGION Network 7: Aborting
   RUNG wire#powerrail
      Contact( "R-202_Write_TO_T-101_DB".Abort )
      Coil( "T-101_Read_FROM_R-202_DB".Aborting )
   END_RUNG
   // the same network as SCL:
   "T-101_Read_FROM_R-202_DB".Aborting := "R-202_Write_TO_T-101_DB".Abort;
END_REGION

REGION Network 8: Release Tank
   RUNG wire#powerrail
      Contact( "R-202_Write_TO_T-101_DB".ReleaseTank )
      Coil( "T-101_Read_FROM_R-202_DB".ReleaseTank )
   END_RUNG
   // the same network as SCL:
   "T-101_Read_FROM_R-202_DB".ReleaseTank := "R-202_Write_TO_T-101_DB".ReleaseTank;
END_REGION
END_FUNCTION

// folder: State MACHINE/1)Tanks/Tank T-101 (X)/T-101 <---> T-104

FUNCTION "T-101_Signals_FROM_T-104" : Void   // FC56, LAD
{ S7_Optimized_Access := 'TRUE' }
VERSION : 0.1
BEGIN

REGION Network 1: Start Sequence
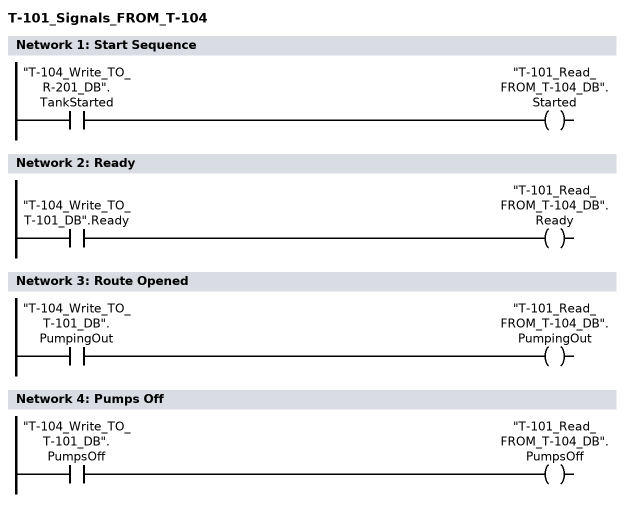
   RUNG wire#powerrail
      Contact( "T-104_Write_TO_R-201_DB".TankStarted )
      Coil( "T-101_Read_FROM_T-104_DB".Started )
   END_RUNG
   // the same network as SCL:
   "T-101_Read_FROM_T-104_DB".Started := "T-104_Write_TO_R-201_DB".TankStarted;
END_REGION

REGION Network 2: Ready
   RUNG wire#powerrail
      Contact( "T-104_Write_TO_T-101_DB".Ready )
      Coil( "T-101_Read_FROM_T-104_DB".Ready )
   END_RUNG
   // the same network as SCL:
   "T-101_Read_FROM_T-104_DB".Ready := "T-104_Write_TO_T-101_DB".Ready;
END_REGION

REGION Network 3: Route Opened
   RUNG wire#powerrail
      Contact( "T-104_Write_TO_T-101_DB".PumpingOut )
      Coil( "T-101_Read_FROM_T-104_DB".PumpingOut )
   END_RUNG
   // the same network as SCL:
   "T-101_Read_FROM_T-104_DB".PumpingOut := "T-104_Write_TO_T-101_DB".PumpingOut;
END_REGION

REGION Network 4: Pumps Off
   RUNG wire#powerrail
      Contact( "T-104_Write_TO_T-101_DB".PumpsOff )
      Coil( "T-101_Read_FROM_T-104_DB".PumpsOff )
   END_RUNG
   // the same network as SCL:
   "T-101_Read_FROM_T-104_DB".PumpsOff := "T-104_Write_TO_T-101_DB".PumpsOff;
END_REGION
END_FUNCTION

// folder: State MACHINE/1)Tanks/Tank T-102 (Y)

FUNCTION_BLOCK "T-102_SEQ"   // FB42, GRAPH_PLUS
{ S7_Optimized_Access := 'TRUE' }